   (* revision history
   hm  21. mar. 2008   rev 1.0
       original version

   hm  10. mar. 2009 rev 1.1
       real constants updated to new systax using dot

   *)
END_FUNCTION

FUNCTION "R2_ADD" : "REAL2"   // FC144, SCL
TITLE = R2_ADD
{ S7_Optimized_Access := 'FALSE' }
AUTHOR : hugo
FAMILY : R2
NAME : ADD
VERSION : 1.0
// R2_add adds a real to a double real which extends the accuracy of a real to twice as many digits
//  
// uses: REAL2 [UDT11]
   VAR_INPUT
      X : "REAL2";
      Y : Real;
   END_VAR
   VAR_TEMP
      temp : Real;
      tR2_ADD : "REAL2";
   END_VAR
BEGIN


   #temp := #X.RX;
   #tR2_ADD.RX := #Y + #X.R1 + #X.RX;
   #tR2_ADD.R1 := #temp - #tR2_ADD.RX + #Y + #X.R1;

   #R2_ADD := #tR2_ADD;

   (* revision history
   hm      20.3.2008   rev 1.0
       original version

   *)
END_FUNCTION

FUNCTION "R2_ADD2" : "REAL2"   // FC145, SCL
TITLE = R2_ADD2
{ S7_Optimized_Access := 'FALSE' }
AUTHOR : hugo
FAMILY : R2
NAME : ADD2
VERSION : 1.0
// R2_add2 adds a double precision real to a double precision real which extends the accuracy of a real to twice as many digits
//  
// uses: REAL2 [UDT11]
   VAR_INPUT
      X : "REAL2";
      Y : "REAL2";
   END_VAR
   VAR_TEMP
      tR2_ADD2 : "REAL2";
   END_VAR
BEGIN


   #tR2_ADD2.R1 := #X.R1 + #Y.R1;
   #tR2_ADD2.RX := #X.RX + #Y.RX;

   #R2_ADD2 := #tR2_ADD2;

   (* revision history
   hm      20.3.2008   rev 1.0
       original version

   *)
END_FUNCTION

FUNCTION "R2_MUL" : "REAL2"   // FC146, SCL
TITLE = R2_MUL
{ S7_Optimized_Access := 'FALSE' }
AUTHOR : hugo
FAMILY : R2
NAME : MUL
VERSION : 1.0
// R2_mul multiplies a real with a double real which extends the accuracy of a real to twice as many digits
//  
// uses: REAL2 [UDT11]
   VAR_INPUT
      X : "REAL2";
      Y : Real;
   END_VAR
   VAR_TEMP
      tR2_MUL : "REAL2";
   END_VAR
BEGIN


   #tR2_MUL.RX := #X.RX * #Y;
   #tR2_MUL.R1 := #X.R1 * #Y;

   #R2_MUL := #tR2_MUL;

   (* revision history
   hm      20.3.2008   rev 1.0
       original version

   *)
END_FUNCTION

FUNCTION "R2_SET" : "REAL2"   // FC147, SCL
TITLE = R2_SET
{ S7_Optimized_Access := 'FALSE' }
AUTHOR : hugo
FAMILY : R2
NAME : SET
VERSION : 1.1
// R2_set sets a double precision real to a single real value.
// 
// uses: REAL2 [UDT11]
   VAR_INPUT
      X : Real;
   END_VAR
   VAR_TEMP
      tR2_SET : "REAL2";
   END_VAR
BEGIN


   #tR2_SET.RX := #X;
   #tR2_SET.R1 := 0.0;

   #R2_SET := #tR2_SET;


   (* revision history
   hm  2. jun. 2008    rev 1.0
       original version

   hm  10. mar. 2009   rev 1.1
       real constants updated to new systax using dot

   *)
END_FUNCTION

// ===== PLC "Math Vektormathematik"  Unspecific CPU S7 300 =====

TYPE "VECTOR_3"
VERSION : 0.0
   STRUCT
      X : Real;
      Y : Real;
      Z : Real;
   END_STRUCT;
END_TYPE

FUNCTION "V3_ABS" : Real   // FC162, SCL
TITLE = V3_ABS
{ S7_Optimized_Access := 'FALSE' }
AUTHOR : hugo
FAMILY : MATH_V3
NAME : V3_ABS
VERSION : 1.0
// this function calculates the length of a vectors in a 3 dimensional space
// 
// uses: VECTOR_3 [UDT15]
   VAR_INPUT
      "A" : "VECTOR_3";
   END_VAR
BEGIN


   #V3_ABS := SQRT(#"A".X * #"A".X + #"A".Y * #"A".Y + #"A".Z * #"A".Z);


   (* revision history
   hm    11 dec 2007 rev 1.0
     original version

   *)
END_FUNCTION

FUNCTION "V3_ADD" : "VECTOR_3"   // FC163, SCL
TITLE = V3_ADD
{ S7_Optimized_Access := 'FALSE' }
AUTHOR : hugo
FAMILY : MATH_V3
NAME : V3_ADD
VERSION : 1.0
// this function adds two vectors in a 3 dimensional space
// 
// uses: VECTOR_3 [UDT15]
   VAR_INPUT
      "A" : "VECTOR_3";
      "B" : "VECTOR_3";
   END_VAR
BEGIN


     #V3_ADD.X := #"A".X + #"B".X;
     #V3_ADD.Y := #"A".Y + #"B".Y;
     #V3_ADD.Z := #"A".Z + #"B".Z;

     #V3_ADD := #V3_ADD;


   (* revision history
   hm    11 dec 2007 rev 1.0
     original version

   *)
END_FUNCTION

FUNCTION "V3_ANG" : Real   // FC164, SCL
TITLE = V3_ANG
{ S7_Optimized_Access := 'FALSE' }
AUTHOR : hugo
FAMILY : MATH_V3
NAME : V3_ANG
VERSION : 1.1
// this function calculates the angle between two vectors in a 3 dimensional space
// 
// uses: VECTOR_3 [UDT15]
//       V3_ABS [FC162]
//       V3_DPRO [FC165]
   VAR_INPUT
      "A" : "VECTOR_3";
      "B" : "VECTOR_3";
   END_VAR
   VAR_TEMP
      d : Real;
      temp_A : "VECTOR_3";
      temp_B : "VECTOR_3";
   END_VAR
BEGIN


   #temp_A := #"A";
   #temp_B := #"B";

   #d := "V3_ABS"(#temp_A) * "V3_ABS"(#temp_B);
   IF #d > 0.0 THEN
       #V3_ANG := ACOS(LIMIT(MN:=-1.0,IN:="V3_DPRO"(A:=#temp_A,B:=#temp_B) / #d,MX:=1.0));
   END_IF;


   (* revision history
   hm  11. dec. 2007   rev 1.0
       original version

   hm  10. mar. 2009   rev 1.1
       changed syntax of real constants to 0.0

   *)
END_FUNCTION

FUNCTION "V3_DPRO" : Real   // FC165, SCL
TITLE = V3_DPRO
{ S7_Optimized_Access := 'FALSE' }
AUTHOR : hugo
FAMILY : MATH_V3
NAME : V3_DPRO
VERSION : 1.0
// this function calculates the dot product of two vectors in 3 dimensional space
// 
// uses: VECTOR_3 [UDT15]
   VAR_INPUT
      "A" : "VECTOR_3";
      "B" : "VECTOR_3";
   END_VAR
BEGIN


     #V3_DPRO := #"A".X * #"B".X + #"A".Y * #"B".Y + #"A".Z * #"B".Z;


   (* revision history
   hm    11 dec 2007 rev 1.0
     original version

   *)
END_FUNCTION

FUNCTION "V3_NORM" : "VECTOR_3"   // FC166, SCL
TITLE = V3_NORM
{ S7_Optimized_Access := 'FALSE' }
AUTHOR : hugo
FAMILY : MATH_V3
NAME : V3_NORM
VERSION : 1.1
// this function generates a vectors with absolute length 1 from a vector A in a 3 dimensional space
// 
// uses: VECTOR_3 [UDT15]
//       V3_ABS [FC162]
//       V3_SMUL [FC170]
   VAR_INPUT
      "A" : "VECTOR_3";
   END_VAR
   VAR_TEMP
      la : Real;
      temp_A : "VECTOR_3";
      temp_V3_NORM : "VECTOR_3";
   END_VAR
BEGIN


   #temp_A := #"A";

   #la := "V3_ABS"(#temp_A);
   IF #la > 0.0 THEN
       #temp_V3_NORM := "V3_SMUL"(A:=#temp_A,M:=1.0 / #la);
   END_IF;

   #V3_NORM := #temp_V3_NORM;


   (* revision history
   hm  11 dec 2007 rev 1.0
       original version

   hm  10. mar. 2009   rev 1.1
       changed syntax of real constants to 0.0

   *)
END_FUNCTION

FUNCTION "V3_NUL" : Bool   // FC167, SCL
TITLE = V3_NUL
{ S7_Optimized_Access := 'FALSE' }
AUTHOR : hugo
FAMILY : MATH_V3
NAME : V3_NUL
VERSION : 1.1
// this function checks if a vectors in a null Vector
// 
// uses: VECTOR_3 [UDT15]
   VAR_INPUT
      "A" : "VECTOR_3";
   END_VAR
BEGIN


   #V3_NUL := #"A".X = 0.0 AND #"A".Y = 0.0 AND #"A".Z = 0.0;


   (* revision history
   hm  12 dec 2007 rev 1.0
       original version

   hm  10. mar. 2009   rev 1.1
       changed syntax of real constants to 0.0

   *)
END_FUNCTION

FUNCTION "V3_PAR" : Bool   // FC168, SCL
TITLE = V3_PAR
{ S7_Optimized_Access := 'FALSE' }
AUTHOR : hugo
FAMILY : MATH_V3
NAME : V3_PAR
VERSION : 1.1
// this function checks if two vectors in a 3 dimensional space are parallel.
// which means the two vectors have the same direction
// 
// uses: VECTOR_3 [UDT15]
//       V3_ABS [FC162]
//       V3_XPRO [FC173]
   VAR_INPUT
      "A" : "VECTOR_3";
      "B" : "VECTOR_3";
   END_VAR
   VAR_TEMP
      temp_A : "VECTOR_3";
      temp_B : "VECTOR_3";
   END_VAR
BEGIN


   #temp_A := #"A";
   #temp_B := #"B";

   #V3_PAR := "V3_ABS"("V3_XPRO"(A:=#temp_A,B:=#temp_B)) = 0.0;


   (* revision history
   hm  11 dec 2007   rev 1.0
       original version

   hm  10. mar. 2009   rev 1.1
       changed syntax of real constants to 0.0

   *)
END_FUNCTION

FUNCTION "V3_REV" : "VECTOR_3"   // FC169, SCL
TITLE = V3_REV
{ S7_Optimized_Access := 'FALSE' }
AUTHOR : hugo
FAMILY : MATH_V3
NAME : V3_REV
VERSION : 1.0
// this function reverses a vector in a 3 dimensional space
// 
// uses: VECTOR_3 [UDT15]
   VAR_INPUT
      "A" : "VECTOR_3";
   END_VAR
   VAR_TEMP
      temp_V3_REV : "VECTOR_3";
   END_VAR
BEGIN


     #temp_V3_REV.X := -#"A".X;
     #temp_V3_REV.Y := -#"A".Y;
     #temp_V3_REV.Z := -#"A".Z;

     #V3_REV := #temp_V3_REV;

   (* revision history
   hm    11 dec 2007 rev 1.0
     original version

   *)
END_FUNCTION

FUNCTION "V3_SMUL" : "VECTOR_3"   // FC170, SCL
TITLE = V3_SMUL
{ S7_Optimized_Access := 'FALSE' }
AUTHOR : hugo
FAMILY : MATH_V3
NAME : V3_SMUL
VERSION : 1.0
// this function multiplies a vectors in a 3 dimensional space with a skalar M
// 
// uses: VECTOR_3 [UDT15]
   VAR_INPUT
      "A" : "VECTOR_3";
      "M" : Real;
   END_VAR
   VAR_TEMP
      temp_V3_SMUL : "VECTOR_3";
   END_VAR
BEGIN


   #temp_V3_SMUL.X := #"A".X * #"M";
   #temp_V3_SMUL.Y := #"A".Y * #"M";
   #temp_V3_SMUL.Z := #"A".Z * #"M";

   #V3_SMUL := #temp_V3_SMUL;


   (* revision history
   hm    11 dec 2007 rev 1.0
     original version

   *)
END_FUNCTION

FUNCTION "V3_SUB" : "VECTOR_3"   // FC171, SCL
TITLE = V3_SUB
{ S7_Optimized_Access := 'FALSE' }
AUTHOR : hugo
FAMILY : MATH_V3
NAME : V3_SUB
VERSION : 1.0
// this function subtracts two vectors in a 3 dimensional space
// V3_SUB = A - B
// 
// uses: VECTOR_3 [UDT15]
   VAR_INPUT
      "A" : "VECTOR_3";
      "B" : "VECTOR_3";
   END_VAR
   VAR_TEMP
      temp_V3_SUB : "VECTOR_3";
   END_VAR
BEGIN


     #temp_V3_SUB.X := #"A".X - #"B".X;
     #temp_V3_SUB.Y := #"A".Y - #"B".Y;
     #temp_V3_SUB.Z := #"A".Z - #"B".Z;

     #V3_SUB := #temp_V3_SUB;

   (* revision history
   hm    11 dec 2007 rev 1.0
     original version

   *)
END_FUNCTION

FUNCTION "V3_XANG" : Real   // FC172, SCL
TITLE = V3_XANG
{ S7_Optimized_Access := 'FALSE' }
AUTHOR : hugo
FAMILY : MATH_V3
NAME : V3_XANG
VERSION : 1.1
// this function calculates the angle between the X-axis and a vectors in a 3 dimensional space
// 
// uses: VECTOR_3 [UDT15]
//       V3_ABS [FC162]
   VAR_INPUT
      "A" : "VECTOR_3";
   END_VAR
   VAR_TEMP
      la : Real;
      temp_A : "VECTOR_3";
   END_VAR
BEGIN


   #temp_A := #"A";

   #la := "V3_ABS"(#temp_A);
   IF #la > 0.0 THEN
       #V3_XANG := ACOS(#temp_A.X / #la);
   END_IF;


   (* revision history
   hm  11 dec 2007   rev 1.0
       original version

   hm  10. mar. 2009   rev 1.1
       changed syntax of real constants to 0.0

   *)
END_FUNCTION

FUNCTION "V3_XPRO" : "VECTOR_3"   // FC173, SCL
TITLE = V3_XPRO
{ S7_Optimized_Access := 'FALSE' }
AUTHOR : hugo
FAMILY : MATH_V3
NAME : V3_XPRO
VERSION : 1.0
// this function adds two vectors in a 3 dimensional space
// 
// uses: VECTOR_3 [UDT15]
   VAR_INPUT
      "A" : "VECTOR_3";
      "B" : "VECTOR_3";
   END_VAR
   VAR_TEMP
      temp_V3_XPRO : "VECTOR_3";
   END_VAR
BEGIN


   #temp_V3_XPRO.X := #"A".Y * #"B".Z - #"A".Z * #"B".Y;
   #temp_V3_XPRO.Y := #"A".Z * #"B".X - #"A".X * #"B".Z;
   #temp_V3_XPRO.Z := #"A".X * #"B".Y - #"A".Y * #"B".X;

   #V3_XPRO := #temp_V3_XPRO;

   (* revision history
   hm    11 dec 2007 rev 1.0
     original version

   *)
END_FUNCTION

FUNCTION "V3_YANG" : Real   // FC174, SCL
TITLE = V3_YANG
{ S7_Optimized_Access := 'FALSE' }
AUTHOR : hugo
FAMILY : MATH_V3
NAME : V3_YANG
VERSION : 1.1
// this function calculates the angle between the Y-axis and a vectors in a 3 dimensional space
// 
// uses: VECTOR_3 [UDT15]
//       V3_ABS [FC162]
   VAR_INPUT
      "A" : "VECTOR_3";
   END_VAR
   VAR_TEMP
      la : Real;
      temp_A : "VECTOR_3";
   END_VAR
BEGIN


   #temp_A := #"A";

   #la := "V3_ABS"(#temp_A);
   IF #la > 0.0 THEN
       #V3_YANG := ACOS(#temp_A.Y / #la);
   END_IF;


   (* revision history
   hm  11 dec 2007   rev 1.0
       original version

   hm  10. mar. 2009   rev 1.1
       changed syntax of real constants to 0.0

   *)
END_FUNCTION

FUNCTION "V3_ZANG" : Real   // FC175, SCL
TITLE = V3_ZANG
{ S7_Optimized_Access := 'FALSE' }
AUTHOR : hugo
FAMILY : MATH_V3
NAME : V3_ZANG
VERSION : 1.1
// this function calculates the angle between the Z-axis and a vectors in a 3 dimensional space
// 
// uses: VECTOR_3 [UDT15]
//       V3_ABS [FC162]
   VAR_INPUT
      "A" : "VECTOR_3";
   END_VAR
   VAR_TEMP
      la : Real;
      temp_A : "VECTOR_3";
   END_VAR
BEGIN


   #temp_A := #"A";

   #la := "V3_ABS"(#temp_A);
   IF #la > 0.0 THEN
       #V3_ZANG := ACOS(#temp_A.Z / #la);
   END_IF;


   (* revision history
   hm  11 dec 2007   rev 1.0
       original version

   hm  10. mar. 2009   rev 1.1
       changed syntax of real constants to 0.0

   *)
END_FUNCTION

// ===== PLC "Mathematical"  Unspecific CPU S7 300 =====

VAR_GLOBAL CONSTANT   // PLC tag table "STEP7 classic symbols"
   "PI1" : Real := 3.14159265358979323846264338327950288;
   "PI05" : Real := 1.5707963267949;
   "PI2" : Real := 6.283185307179586476;   // PI * 2
   "E_INV" : Real := 0.367879441171442;   // 1 / e
   "PI_INV" : Real := 0.318309886183791;   // 1 / PI
   "debug" : Bool := FALSE;
   "N" : Int := 0;
   "offset" : Int := 0;
   "E" : Real := 2.71828182845904523536028747135266249;   // Eulersche Konstante
   "PI" : Real := 3.14159265358979323846264338327950288;
   "offset_1" : DWord := 0;
END_VAR

TYPE "FRACTION"
VERSION : 0.0
   STRUCT
      NUMERATOR : Int;
      DENOMINATOR : Int;
   END_STRUCT;
END_TYPE

DATA_BLOCK "MATH"   // DB2
TITLE = MATH
{ S7_Optimized_Access := 'FALSE' }
AUTHOR : oscat
FAMILY : CONSTANT
NAME : DBMATH
VERSION : 1.1
   VAR
      PI : Real := 3.141593e+0;   // Kreiszahl PI
      PI2 : Real := 6.283185e+0;   // PI * 2
      PI4 : Real := 1.256637e+1;   // PI * 4
      PI05 : Real := 1.570796e+0;   // PI / 2
      PI025 : Real := 7.853982e-1;   // PI / 4
      PI_INV : Real := 3.183099e-1;   // 1 / PI
      "E" : Real := 2.718282e+0;   // Eulersche Konstante
      E_INV : Real := 3.678795e-1;   // 1 / e
      SQ2 : Real := 1.414214e+0;   // Wurzel von 2
      FACTS : Array[0..12] of DInt;
   END_VAR
BEGIN
   FACTS[0] := DINT#1;
   FACTS[1] := DINT#1;
   FACTS[2] := DINT#2;
   FACTS[3] := DINT#6;
   FACTS[4] := DINT#24;
   FACTS[5] := DINT#120;
   FACTS[6] := DINT#720;
   FACTS[7] := DINT#5040;
   FACTS[8] := DINT#40320;
   FACTS[9] := DINT#362880;
   FACTS[10] := DINT#3628800;
   FACTS[11] := DINT#39916800;
   FACTS[12] := DINT#479001600;
END_DATA_BLOCK

DATA_BLOCK "IDB_STIME"   // DB64
{ S7_Optimized_Access := 'FALSE' }
AUTHOR : dalbi
FAMILY : MEASURE
VERSION : 0.0
// stored: InstanceOfName STIME
"STIME"
BEGIN
END_DATA_BLOCK

FUNCTION_BLOCK "STIME"   // FB64, SCL
TITLE = STIME
{ S7_Optimized_Access := 'FALSE' }
AUTHOR : dalbi
FAMILY : MEASURE
NAME : STIME
VERSION : 1.4
// this function block makes sure that the timer of a siemens sps counts from 0 - 2^32-1.
   VAR_OUTPUT
      tx : DWord;
      at_tx AT tx : Array[0..31] of Bool;
   END_VAR
   VAR
      last_time : DWord;
      bit31 : Bool;
      init : Bool := TRUE;
   END_VAR
   VAR_TEMP
      TOP_SI : Struct
         EV_CLASS : Byte;
         EV_NUM : Byte;
         PRIORITY : Byte;
         NUM : Byte;
         TYP2_3 : Byte;
         TYP1 : Byte;
         ZI1 : Word;
         ZI2_3 : DWord;
      END_STRUCT;
      START_UP_SI : Struct
         EV_CLASS : Byte;
         EV_NUM : Byte;
         PRIORITY : Byte;
         NUM : Byte;
         TYP2_3 : Byte;
         TYP1 : Byte;
         ZI1 : Word;
         ZI2_3 : DWord;
      END_STRUCT;
      ERR : Int;
   END_VAR
BEGIN


   (* this FB is only necessary for siemens sps
   the siemens sps timer counts from 0 to 2^31-1 and starts at 0 sfter overrun.
   this means that the bit 31 (the highest bit ) will never be used and therefore
   a problem arises when t2 - t1 is checked.
   t2 - t1 is always valid also in an timer overrun situation where the time t1 is very high and t2 is very low.
   the result of the subtraction t2 - t1 however is still valid.
   this calculation does not work for soiemens because the highest bit is not used.

   this module stores the highest bit, changes the highest bit at every overrun occurence and stuffs ther highest bit in the output.
   the output is then used by t_plc_us and t_plc_ms.

   the correction needs and fb and not a function because the value of the highest bit has to be stored.

   do never use this function block in a codesys environment. the timer in codesys is correct and runs from 0 to 2^32-1
   *)

   (* read actual startup info *)
   (* OB1_SCAN_1  BYTE  -  B#16#01: Abschluss des Neustarts (Warmstarts)
                        -  B#16#02: Abschluss des Wiederanlaufs
                        -  B#16#03: Abschluss des freien Zyklus
                        -  B#16#04: Abschluss des Kaltstarts
                        -  B#16#05: Erster OB 1-Zyklus der neuen Master-CPU nach 
                                    Master-Reserve-Umschaltung und STOP des 
                                    bisherigen Masters *)

   #ERR := RD_SINFO (TOP_SI => #TOP_SI, START_UP_SI => #START_UP_SI);

   (* reset last_time on system startup *)
   IF #TOP_SI.EV_NUM = 1 OR #TOP_SI.EV_NUM = 2 OR #TOP_SI.EV_NUM = 4 OR NOT #init THEN 
       #last_time := 0;
       #bit31 := false;
       #init := true;
   END_IF;

   (* read the system timer *)
   #tx := DINT_TO_DWORD(T_CONV(TIME_TCK()));

   (* check for overrun *)
   IF DWORD_TO_DINT(#tx) < DWORD_TO_DINT(#last_time) THEN
       (* an overrun has occured, change the value of the highest bit *)
       #bit31 := NOT #bit31;
   END_IF;

   (* stuff the highest bit into the timer value *)
   #at_tx[7] := #bit31;

   (* remember the last system time for the next overrun check *)
   #last_time := #tx;


   (* revision history
   DA  14.9.2007 rev 1.0
     original version

   DA  24.2.2008 rev 1.1
     added self reset on system startup

   DA   2.5.2008 rev 1.2
     corect a problem running under OB35

   DA  12.3.2009 rev 1.3
     corect a problem run on different CPUs

   DA  22.12.2009 rev 1.4
     corect a problem on startup
   *)
END_FUNCTION_BLOCK

FUNCTION "DEC1" : Int   // FC52, SCL
TITLE = DEC1
{ S7_Optimized_Access := 'FALSE' }
AUTHOR : hugo
FAMILY : MATH
NAME : DEC1
VERSION : 1.1
// This is a decrement function which decrements the variable X by 1 and if 0 is reached, it begins with M again.
// _dec1(3,X) will generate 3,2,1,0,3,2,...
   VAR_INPUT
      X : Int;
      N : Int;
   END_VAR
BEGIN


   IF #X = 0 THEN
       #DEC1 := #N - 1;
   ELSE
       #DEC1 := #X - 1;
   END_IF;

   (* this is a very elegant version but 50% slower
   X := (X - 1 + N) MOD N;
   *)


   (* revision history
   hm  13. oct. 2008   rev 1.0
       original version

   hm  27. oct. 2008   rev 1.1
       added statement to return value for compatibility reasons
   *)
END_FUNCTION

FUNCTION "INC1" : Int   // FC53, SCL
TITLE = INC1
{ S7_Optimized_Access := 'FALSE' }
AUTHOR : hugo
FAMILY : MATH
NAME : INC1
VERSION : 1.2
// This is a increment function which increments the variable X by 1 and if M is reached, it begins with 0 again.
// _inc1(3,X) will generate 0,1,2,3,0,1,.....
   VAR_INPUT
      X : Int;
      N : Int;
   END_VAR
BEGIN


   IF #X >= #N - 1 THEN
       #INC1 := 0;
   ELSE
       #INC1 := #X + 1;
   END_IF;


   (* this elegant version is 50% slower
   INC1 := X := (x + 1) MOD N;
   *)



   (* revision history
   hm  13. oct. 2008   rev 1.0
       original version

   hm  22. oct. 2008   rev 1.1
       added statement to return value for compatibility reasons

   hm  23. feb. 2009   rev 1.2
       when inc1 is called with X >= N inc will continue with 0
   *)
END_FUNCTION

FUNCTION "ACOSH" : Real   // FC54, SCL
TITLE = ACOSH
{ S7_Optimized_Access := 'FALSE' }
AUTHOR : hugo
FAMILY : MATH
NAME : ACOSH
VERSION : 1.3
// this function calculates the arcus cos hyperbolicus
   VAR_INPUT
      X : Real;
   END_VAR
BEGIN



   #ACOSH := LN(SQRT(#X * #X - 1.0) + #X);


   (* revision history
   hm      12 jan 2007 rev 1.0
       original version

   hm      2. dec 2007 rev 1.1
       changed code for better performance

   hm  16. mar. 2007       rev 1.2
       changed sequence of calculations to improve performance

   hm  10. mar. 2009       rev 1.3
       real constants updated to new systax using dot

   *)
END_FUNCTION

FUNCTION "ACOTH" : Real   // FC55, SCL
TITLE = ACOTH
{ S7_Optimized_Access := 'FALSE' }
AUTHOR : hugo
FAMILY : MATH
NAME : ACOTH
VERSION : 1.2
// this function calculates the arcus cotangens hyperbolicus
   VAR_INPUT
      X : Real;
   END_VAR
BEGIN


   #ACOTH := LN((#X+1.0)/(#X-1.0))*0.5;


   (* revision history
   hm      12 jan 2007 rev 1.0
       original version

   hm      5. jan 2008 rev 1.1
       improved code for better performance

   hm  10. mar. 2009       rev 1.2
       real constants updated to new systax using dot

   *)
END_FUNCTION

FUNCTION "AGDF" : Real   // FC56, SCL
TITLE = AGDF
{ S7_Optimized_Access := 'FALSE' }
AUTHOR : hugo
FAMILY : MATH
NAME : AGDF
VERSION : 1.1
// this function calculates the inverse Gudermannian function.
   VAR_INPUT
      X : Real;
   END_VAR
BEGIN


   #AGDF := LN((1.0 + SIN(#X))/COS(#X));

   (* comment
   the current implementation gives sufficient accuracy only up to X = 1.57 or an output > 10.
   is X closer to PI/2 then the function is more and more unreliable
   *)


   (* revision history
   hm  27. apr. 2008   rev 1.0
       original version

   hm  10. mar. 2009   rev 1.1
       real constants updated to new systax using dot

   *)
END_FUNCTION

FUNCTION "ASINH" : Real   // FC57, SCL
TITLE = ASINH
{ S7_Optimized_Access := 'FALSE' }
AUTHOR : hugo
FAMILY : MATH
NAME : ASINH
VERSION : 1.3
// this function calculates the arcus sin hyperbolicus
   VAR_INPUT
      X : Real;
   END_VAR
BEGIN


   #ASINH := LN(SQRT(#X * #X + 1.0)+#X);


   (* revision history
   hm      12 jan 2007 rev 1.0
       original version

   hm      2. dec 2007 rev 1.1
       changed code for better performance

   hm      16.3. 2007      rev 1.2
       changed sequence of calculations to improve performance

   hm  10. mar. 2009       rev 1.3
       real constants updated to new systax using dot

   *)
END_FUNCTION

FUNCTION "ATAN2" : Real   // FC58, SCL
TITLE = ATAN2
{ S7_Optimized_Access := 'FALSE' }
AUTHOR : hugo
FAMILY : MATH
NAME : ATAN2
VERSION : 1.2
// this function calculates the angle in a coordinate system in rad.
   VAR_INPUT
      Y : Real;
      X : Real;
   END_VAR
BEGIN


   IF #X > 0.0 THEN
       #ATAN2 := ATAN(#Y/#X);
   ELSIF #X < 0.0 THEN
       IF #Y >= 0.0 THEN
           #ATAN2 := ATAN(#Y/#X) + "PI1";
       ELSE
           #ATAN2 := ATAN(#Y/#X) - "PI1";
       END_IF;
   ELSIF #Y > 0.0 THEN
       #ATAN2 := "PI05";
   ELSIF #Y < 0.0 THEN
       #ATAN2 := -"PI05";
   ELSE
       #ATAN2 := 0.0;
   END_IF;


   (* revision history
   hm  20.  apr. 2008  rev 1.0
       original version

   hm  18. oct. 2008   rev 1.1
       changed to use math constants

   hm  10. mar. 2009   rev 1.2
       real constants updated to new systax using dot

   *)
END_FUNCTION

FUNCTION "ATANH" : Real   // FC59, SCL
TITLE = ATANH
{ S7_Optimized_Access := 'FALSE' }
AUTHOR : hugo
FAMILY : MATH
NAME : ATANH
VERSION : 1.2
// this function calculates the arcus tangens hyperbolicus
   VAR_INPUT
      X : Real;
   END_VAR
BEGIN


   #ATANH := LN((1.0 + #X)/(1.0 - #X)) * 0.5;

   (* revision history
   hm      12 jan 2007 rev 1.0
       original version

   hm      5. jan 2008 rev 1.1
       improved code for better performance

   hm  10. mar. 2009     rev 1.2
       real constants updated to new systax using dot

   *)
END_FUNCTION

FUNCTION "BETA" : Real   // FC60, SCL
TITLE = BETA
{ S7_Optimized_Access := 'FALSE' }
AUTHOR : hugo
FAMILY : MATH
NAME : BETA
VERSION : 1.0
// this function calculates the beta function for real number > 0.
// 
// uses: GAMMA [FC84]
   VAR_INPUT
      X : Real;
      Y : Real;
   END_VAR
BEGIN


   #BETA := "GAMMA"(#X) * "GAMMA"(#Y) / "GAMMA"(#X + #Y);


   (* revision history
   hm  26. oct. 2008   rev 1.0
       original version

   *)
END_FUNCTION

FUNCTION "BINOM" : DInt   // FC61, SCL
TITLE = BINOM
{ S7_Optimized_Access := 'FALSE' }
AUTHOR : hugo
FAMILY : MATH
NAME : BINOM
VERSION : 1.0
// this FUNCTION calculates the binomialkoefficient (N over k)
   VAR_INPUT
      N : Int;
      K : Int;
   END_VAR
   VAR_TEMP
      i : Int;
      tK : Int;
      tn : Int;
   END_VAR
BEGIN


   #tK := #K;
   #tn := #N;

   IF 2 * #tK > #tn THEN
       #tK := #tn - #tK;
   END_IF;
   IF #tK > #tn THEN
       RETURN;
   ELSIF #tK = 0 OR #tK = #tn THEN
       #BINOM := 1;
   ELSIF #tK = 1 THEN
       #BINOM := #tn;
   ELSE
       #BINOM := #tn;
       #tn := #tn + 1;
       FOR #i := 2 TO #tK DO
           #BINOM := #BINOM * (#tn - #i) / #i;
       END_FOR;
   END_IF;



   (*
   binomialkoeffizient(n, k)
   1  wenn k = 0 return 1
   2  wenn 2k > n
   3      dann führe aus ergebnis \leftarrow binomialkoeffizient(n, n-k)
   4  sonst führe aus ergebnis \leftarrow n
   5          von i \leftarrow 2 bis k
   6              führe aus ergebnis \leftarrow ergebnis \cdot (n + 1 - i)
   7                        ergebnis \leftarrow ergebnis : i
   8  return ergebnis
   *)



   (* revision history
   hm  25. oct. 2008 rev 1.0
       original version


   *)
END_FUNCTION

FUNCTION "CAUCHY" : Real   // FC62, SCL
TITLE = CAUCHY
{ S7_Optimized_Access := 'FALSE' }
AUTHOR : hugo
FAMILY : MATH
NAME : CAUCHY
VERSION : 1.0
// this function calculates the Cauchy distribution function
   VAR_INPUT
      X : Real;
      T : Real;
      U : Real;
   END_VAR
   VAR_TEMP
      tmp : Real;
   END_VAR
BEGIN


   #tmp := #X - #T;
   #CAUCHY := "PI_INV" * #U / (#U*#U + #tmp*#tmp);



   (* revision hisdtory
   hm  26. oct. 2008   rev 1.0
       original version

   *)
END_FUNCTION

FUNCTION "CAUCHYCD" : Real   // FC63, SCL
TITLE = CAUCHYCD
{ S7_Optimized_Access := 'FALSE' }
AUTHOR : hugo
FAMILY : MATH
NAME : CAUCHYCD
VERSION : 1.0
// this function calculates the Cauchy distribution function
   VAR_INPUT
      X : Real;
      T : Real;
      U : Real;
   END_VAR
BEGIN


   #CAUCHYCD := 0.5 + "PI_INV" * ATAN((#X - #T) / #U);



   (* revision hisdtory
   hm  26. oct. 2008   rev 1.0
       original version

   *)
END_FUNCTION

FUNCTION "T_PLC_MS" : DWord   // FC64, SCL
TITLE = T_PLC_MS
{ S7_Optimized_Access := 'FALSE' }
AUTHOR : hugo
FAMILY : MEASURE
NAME : T_PLC_MS
VERSION : 1.2
// T_PLC_MS reads the internal PLC timer and return the time, it has the advantage to be able to set a debug mode 
// and speed up the counter to test the plc timer overrun which occurs every 50 days respectively 25 days at siemens S7
// this routine also allows to correct the behavior of s7 where the internal plc counter will not count all 32 bits.
// 
// uses: STIME [FB64],IDB_STIME [DB64]
BEGIN


   "IDB_STIME"(); 
   #T_PLC_MS := "IDB_STIME".tx; 
   (* hier muss die korrektur für step7 stattfinden
   plctime muss den vollen wertebereich von time ausnutzen:
   wenn bei step7 time -24tage bis plus 24 tage ist dann muss der timer auch beim überlauf auf -24tage springen 
   und auf keinen fall auf 0 !!!!
   für siemens muss ein weiterer fb im main eingebunden werden der sicherstellt das alle 32 bits durchgezählt werden.
   es kann nur ein fb sein den er muss sich das oberste (32te) bit merken.
   oder etwa spring s7 bei überlauf auf -24 tage????? dann wäre keine korrektur nötig.
   *)
   IF "debug" THEN
       #T_PLC_MS := DINT_TO_DWORD((DWORD_TO_DINT(SHL(IN:=#T_PLC_MS,N:="N") OR SHL(IN:=DWORD#1,N:="N"))-1) + DWORD_TO_DINT("offset_1"));
   END_IF;


   (* revision history
   hm  14.9.2007   rev 1.0
       original version

   hm  12. nov 2007    rev 1.1
       added temporaray variable tx because some compilers could not handle time() as an argument

   hm  16. nov. 2008   rev 1.2
       initialized constants with 0 for compatibility reasons
   *)
END_FUNCTION

FUNCTION "CEIL" : Int   // FC66, SCL
TITLE = CEIL
{ S7_Optimized_Access := 'FALSE' }
AUTHOR : hugo
FAMILY : MATH
NAME : CEIL
VERSION : 1.1
// This is a rounding function which returns the smallest possible integer which is greater or equal to X.
// ceil(3.14) = 4
// ceil(-3.14) = 3
   VAR_INPUT
      X : Real;
   END_VAR
BEGIN


     #CEIL := REAL_TO_INT(#X); //DINT_TO_INT(TRUNC(X));
     IF #CEIL < #X THEN
         #CEIL := #CEIL + 1;
     END_IF;

   (* code before rev 1.1
   CEIL := D_TRUNC(X);
   IF CEIL < X THEN
     ceil := ceil + 1;
   END_IF;
   *)

   (* revision history
   hm    7. feb. 2007  rev 1.0
     original version

   hm    21. mar. 2008 rev 1.1
     use REAL_TO_INT instead of trunc for compatibility reasons

   *)
END_FUNCTION

FUNCTION "CEIL2" : DInt   // FC67, SCL
TITLE = CEIL2
{ S7_Optimized_Access := 'FALSE' }
AUTHOR : hugo
FAMILY : MATH
NAME : CEIL
VERSION : 1.3
// This is a rounding function which returns the smallest possible integer which is greater or equal to X.
// ceil2(3.14) = 4
// ceil2(-3.14) = -3
   VAR_INPUT
      X : Real;
   END_VAR
BEGIN


   #CEIL2 := REAL_TO_DINT(#X);
   IF DINT_TO_REAL(#CEIL2) < #X THEN
           #CEIL2 := #CEIL2 + 1;
   END_IF;


   (* revision history
   hm  21. mar. 2008   rev 1.0
       original version

   hm  4. apr. 2008    rev 1.1
       added type conversion to avoid warnings under codesys 3.0

   hm  30. jun. 2008   rev 1.2
       added type conversion to avoid warnings under codesys 3.0

   hm  10. mar. 2009   rev 1.3
       use correct statement real_to_DINT

   *)
END_FUNCTION

FUNCTION "CMP" : Bool   // FC68, SCL
TITLE = CMP
{ S7_Optimized_Access := 'FALSE' }
AUTHOR : hugo
FAMILY : MATH
NAME : CMP
VERSION : 1.1
// this function checks two inputs x and y if they are identical with the first N digits
// example : cmp(3.141516,3.141517,6 is true.
// 
// uses: EXP10 [FC77]
//       FLOOR [FC81]
   VAR_INPUT
      X : Real;
      Y : Real;
      N : Int;
   END_VAR
   VAR_TEMP
      tmp : Real;
   END_VAR
BEGIN


   #tmp := ABS(#X);
   IF #tmp > 0.0 THEN
       #tmp := "EXP10"(INT_TO_REAL("FLOOR"((LN(#tmp)/LN(10)))-#N+1));
   ELSE
       #tmp := "EXP10"(#tmp);
   END_IF;
   #CMP := ABS(#X - #Y) < #tmp;


   (* revision history
   hm  12. mar. 2008   rev 1.0
       original version

   hm  10. mar. 2009   rev 1.1
       added type conversion for compatibility reasons
   *)
END_FUNCTION

FUNCTION "COSH" : Real   // FC69, SCL
TITLE = COSH
{ S7_Optimized_Access := 'FALSE' }
AUTHOR : hugo
FAMILY : MATH
NAME : COSH
VERSION : 1.3
// this function calculates the cos hyperbolicus
   VAR_INPUT
      X : Real;
   END_VAR
   VAR_TEMP
      t : Real;
   END_VAR
BEGIN


   #t := EXP(#X);
   #COSH := (1.0 / #t + #t) * 0.5;


   (* revision histroy
   hm  12.1.2007   rev 1.0
       original version

   hm  1.12.2007   rev 1.1
       changed code to improve performance

   hm  5. jan 2008   rev 1.2
       further performance improvement

   hm  10. mar. 2009   rev 1.3
       real constants updated to new systax using dot
   *)
END_FUNCTION

FUNCTION "COTH" : Real   // FC70, SCL
TITLE = COTH
{ S7_Optimized_Access := 'FALSE' }
AUTHOR : hugo
FAMILY : MATH
NAME : COTH
VERSION : 1.4
// this function calculates the cotangens hyperbolicus
   VAR_INPUT
      X : Real;
   END_VAR
BEGIN


   IF #X > 20.0 THEN
       #COTH :=1.0;
   ELSIF #X < -20.0 THEN
       #COTH := -1.0;
   ELSE
       #COTH := 1.0 + 2.0 / (EXP(#X * 2.0) - 1.0);
   END_IF;


   (* revision histroy
   hm      12.1.2007   rev 1.0
       original version

   hm  1.12.2007       rev 1.1
       changed code to improve performance

   hm  8. jan 2008 rev 1.2
       further improvement in performance

   hm  10. mar 2008    rev 1.3
       extended range of valid inputs to +/- INV
       changed formula for better accuracy

   hm  10. mar. 2009   rev 1.4
       real constants updated to new systax using dot
   *)
END_FUNCTION

FUNCTION "D_TRUNC" : DInt   // FC71, SCL
TITLE = D_TRUNC
{ S7_Optimized_Access := 'FALSE' }
AUTHOR : hugo
FAMILY : MATH
NAME : DTRUNC
VERSION : 1.2
// d_trunc truncates a real to a dint 1.5 will be 1 and -1.5 will be -1
// d_trunc is necessary because many systems do not offer a trunc to a dint
   VAR_INPUT
      X : Real;
   END_VAR
BEGIN


   #D_TRUNC := REAL_TO_DINT(#X);
   IF #X > 0.0 THEN
       IF DINT_TO_REAL(#D_TRUNC) > #X THEN #D_TRUNC := #D_TRUNC - 1; END_IF;
   ELSE
       IF DINT_TO_REAL(#D_TRUNC) < #X THEN #D_TRUNC := #D_TRUNC + 1; END_IF;
   END_IF;


   (* for systems that support a dint truncation this routine can be replaced by trunc() *)


   (* revision history
   hm  21. mar. 2008   rev 1.0
       original version

   hm  31. oct. 2008   rev 1.1
       optimized performance

   hm  10. mar. 2009   rev 1.2
       real constants updated to new systax using dot
   *)
END_FUNCTION

FUNCTION "DEG" : Real   // FC72, SCL
TITLE = DEG
{ S7_Optimized_Access := 'FALSE' }
AUTHOR : hugo
FAMILY : MATH
NAME : DEG
VERSION : 1.2
// this function converts degrees into Radiant
// 
// uses: MODR [FC97]
//       FLOOR2 [FC82]
   VAR_INPUT
      rad : Real;
   END_VAR
BEGIN


   #DEG := "MODR"(IN:=57.29577951308232 * #rad,DIVI:=360.0);


   (* revision history
   hm  4. aug 2006 rev 1.0
       original version

   hm 16. oct 2007 rev 1.1
       added modr statement which prohibits deg to become bigger than 360

   hm  10. mar. 2009   rev 1.2
       real constants updated to new systax using dot
   *)
END_FUNCTION

FUNCTION "DIFFER" : Bool   // FC73, SCL
TITLE = DIFFER
{ S7_Optimized_Access := 'FALSE' }
AUTHOR : hugo
FAMILY : MATH
NAME : DIFFER
VERSION : 1.1
// this function checks if in1 differs more then x from in2
// the output is true if in1 < in2 - x or in1 > in2 + X
   VAR_INPUT
      in1 : Real;
      in2 : Real;
      X : Real;
   END_VAR
BEGIN


   #DIFFER := ABS(#in1 - #in2) > #X;

   (* revision history
   hm    8. oct 2006   rev 1.0
     original version

   hm    16. mar 2008  rev 1.1
     improverd code for performance

   *)
END_FUNCTION

FUNCTION "ERF" : Real   // FC74, SCL
TITLE = ERF
{ S7_Optimized_Access := 'FALSE' }
AUTHOR : hugo
FAMILY : MATH
NAME : ERF
VERSION : 1.3
// this function calculates the erf (error) function.
// 
// uses: SGN [FC106]
   VAR_INPUT
      X : Real;
   END_VAR
   VAR_TEMP
      x2 : Real;
      ax2 : Real;
   END_VAR
BEGIN


   #x2 := #X*#X;
   #ax2 := 0.147 * #x2 + 1.0;
   #ERF := SQRT(1.0 - EXP(-#x2 * ((0.27323954473516 + #ax2)/(#ax2)))) * "SGN"(#X);


   (* revision history
   hm  7. apr. 2008    rev 1.0
       original version

   hm  30. jun. 2008   rev 1.1
       added type conversions to avoid warnings under codesys 3.0

   hm  25. oct. 2008   rev 1.2
       new code using new algorithm

   hm  10. mar. 2009   rev 1.3
       real constants updated to new systax using dot
   *)
END_FUNCTION

FUNCTION "ERFC" : Real   // FC75, SCL
TITLE = ERFC
{ S7_Optimized_Access := 'FALSE' }
AUTHOR : hugo
FAMILY : MATH
NAME : ERFC
VERSION : 1.1
// this function calculates the inverse erf (error) function.
// 
// uses: ERF [FC74]
//       SGN [FC106]
   VAR_INPUT
      X : Real;
   END_VAR
BEGIN


   #ERFC := 1.0 - "ERF"(#X);


   (* revision history
   hm  7. apr. 2008    rev 1.0
       original version

   hm  10. mar. 2009   rev 1.1
       real constants updated to new systax using dot

   *)
END_FUNCTION

FUNCTION "EVEN" : Bool   // FC76, SCL
TITLE = EVEN
{ S7_Optimized_Access := 'FALSE' }
AUTHOR : hugo
FAMILY : MATH
NAME : EVEN
VERSION : 1.2
// this function chacks an input for even value
// the output is true if the input is even.
   VAR_INPUT
      in : DInt;
   END_VAR
   VAR_TEMP
      tIN : DInt;
      _IN AT tIN : Array[0..31] of Bool;
   END_VAR
BEGIN


   #tIN := #in;
   #EVEN := NOT #_IN[24]; //EVEN := NOT in.0;

   (* revision history
   hm  1. oct 2006 rev 1.0
     ORIGINAL VERSION

   hm  01.12.2007  rev 1.1
     changed code for improved performance

   hm  21. mar. 2008 rev 1.2
     changed type of input IN from INT to DINT
   *)
END_FUNCTION

FUNCTION "EXP10" : Real   // FC77, SCL
TITLE = EXP10
{ S7_Optimized_Access := 'FALSE' }
AUTHOR : hugo
FAMILY : MATH
NAME : exp10
VERSION : 1.0
// this function calculates the exponent to the basis 10
// exp10(3) = 1000
   VAR_INPUT
      X : Real;
   END_VAR
BEGIN


     #EXP10 := EXP(#X * 2.30258509299405);

   (* revision history
   hm  2. dec 2007    rev 1.0
     original version

   *)
END_FUNCTION

FUNCTION "EXPN" : Real   // FC78, SCL
TITLE = EXPN
{ S7_Optimized_Access := 'FALSE' }
AUTHOR : hugo
FAMILY : MATH
NAME : EXPN
VERSION : 1.2
// this function calculates X to the power of N (Y = X^N) whilke N is an integer
// especially on CPU's without a floating point unit this algorythm is about 30 times faster then the IEC standard EXPT() Function
   VAR_INPUT
      X : Real;
      N : Int;
   END_VAR
   VAR_TEMP
      tempN : Int;
      _tempN AT tempN : Array[0..15] of Bool;
      tempX : Real;
      sign : Bool;
   END_VAR
BEGIN


   #tempN := #N;
   #tempX := #X;

   #sign := #_tempN[7]; //N.15
   #tempN := ABS(#tempN);
   IF #_tempN[8] THEN #EXPN := #tempX; ELSE #EXPN := 1.0; END_IF;
   #tempN := WORD_TO_INT(SHR(IN:=INT_TO_WORD(#tempN),N:=1));
   WHILE #tempN > 0 DO
      #tempX := #tempX * #tempX;
      IF #_tempN[8] THEN #EXPN := #EXPN * #tempX; END_IF;
      #tempN := WORD_TO_INT(SHR(IN:=INT_TO_WORD(#tempN),N:=1));
   END_WHILE;
   IF #sign THEN #EXPN := 1.0 / #EXPN; END_IF;


   (* revision history
   hm  4. dec 2007 rev 1.0
       original version

   hm  22. oct. 2008   rev 1.1
       optimized code

   hm  10. mar. 2009   rev 1.2
       removed nested comments
       real constants updated to new systax using dot

   *)
END_FUNCTION

FUNCTION "FACT" : DInt   // FC79, SCL
TITLE = FACT
{ S7_Optimized_Access := 'FALSE' }
AUTHOR : hugo
FAMILY : MATH
NAME : FACT
VERSION : 1.5
// this function calculates the factorial of x
// if the input is negative or higher then 12 the output will be -1.
// 
// uses: MATH [DB2]
   VAR_INPUT
      X : Int;
   END_VAR
BEGIN


   IF #X >= 0 AND #X <= 12 THEN
     #FACT := "MATH".FACTS[#X];
   ELSE
     #FACT := -1;
   END_IF;


   (* working code without array
   IF X > 12 OR X < 0 THEN
     FACT := -1;
   ELSIF X < 7 THEN
     FACT := 1;
     FOR i := 2 TO X DO
       FACT := FACT * i;
     END_FOR;
   ELSE
     FACT := 5040;
     FOR i := 8 TO X DO
       FACT := FACT * i;
     END_FOR;
   END_IF;
   *)

   (* revision history
   hm 4.3.2007   rev 1.1
     changed a critical error where while loop was indefinite.

   hm  10.12.2007  rev 1.2
     start value for i has changed to 2 for better performance

   hm  10. mar 2008  rev 1.3
     changed output of fact to dint to allow bigger values

   hm  27. oct. 2008 rev 1.4
     optimized code

   hm  26. mar. 2011 rev 1.5
     using array math.facts
   *)
END_FUNCTION

FUNCTION "FIB" : Real   // FC80, SCL
TITLE = FIB
{ S7_Optimized_Access := 'FALSE' }
AUTHOR : hugo
FAMILY : MATH
NAME : FIB
VERSION : 1.3
// this function calculates the fibonacci sequence
   VAR_INPUT
      X : Int;
   END_VAR
   VAR_TEMP
      tX : Real;
      t_1 : Real;
      t_2 : Real;
   END_VAR
BEGIN


   #t_1 := 0;
   #t_2 := 0;

   #tX := INT_TO_REAL(#X);

   IF #tX < 0 OR #tX > 46 THEN
       #FIB := -1;
   ELSIF #X < 2 THEN
       #FIB := #tX;
       RETURN;
   ELSE
       (* the fibonacci number is the sum of the two suceeding fibonaci numbers *)
       (* we store the numbers alternatively in t1 and t2 depending on pt *)
       #t_2 := 1;
       WHILE #tX > 3 DO
           #tX := #tX-2;
           #t_1 := #t_1 + #t_2;
           #t_2 := #t_1 + #t_2;
       END_WHILE;
       IF #tX > 2 THEN #t_1 := #t_1 + #t_2; END_IF;
       #FIB := #t_1 + #t_2;
   END_IF;

   (* alternative code for very big numbers

   IF X < 31 THEN
       fib := 0.4472136 * (expn(1.618034,X) - expn(-0.618034,X));
   ELSE
       fib := 0.4472133 * expn(1.618034,X);
   END_IF;

   *)

   (* revision history
   hm      27. dec 2007    rev 1.0
       original version

   hm      2. jan 2008 rev 1.1
       deleted unused variable pt

   hm      10. mar 2008    rev 1.2
       changed output to dint instead of real

   hm      26. mar. 2008   rev 1.3
       function now returns -1 for input < 0 or > 46

   *)
END_FUNCTION

FUNCTION "FLOOR" : Int   // FC81, SCL
TITLE = FLOOR
{ S7_Optimized_Access := 'FALSE' }
AUTHOR : hugo
FAMILY : MATH
NAME : FLOOR
VERSION : 1.1
// This is a rounding function which returns the biggest possible integer which is less or equal to X.
// floor(3.14) = 3
// floor(-3.14) = 4
   VAR_INPUT
      X : Real;
   END_VAR
BEGIN


   #FLOOR := REAL_TO_INT(#X);
   IF #FLOOR > #X THEN
       #FLOOR := #FLOOR - 1;
   END_IF;

   (* revision history
   hm    7. feb 2007   rev 1.0
     originlal version

   hm    21. mar. 2008 rev 1.1
     replaced trunc with real_to_int for compatibility reasons

   *)
END_FUNCTION

FUNCTION "FLOOR2" : DInt   // FC82, SCL
TITLE = FLOOR2
{ S7_Optimized_Access := 'FALSE' }
AUTHOR : hugo
FAMILY : MATH
NAME : FLOOR2
VERSION : 1.1
// This is a rounding function which returns the biggest possible integer which is less or equal to X.
// floor2(3.14) = 3
// floor2(-3.14) = -4
   VAR_INPUT
      X : Real;
   END_VAR
BEGIN


   #FLOOR2 := REAL_TO_DINT(#X);
   IF DINT_TO_REAL(#FLOOR2) > #X THEN
     #FLOOR2 := #FLOOR2 - 1;
   END_IF;

   (* revision history
   hm  21. mar. 2008   rev 1.0
       originlal version

   hm  4. apr. 2008    rev 1.1
       added type conversion to avoid warnings under codesys 3.0
   *)
END_FUNCTION

FUNCTION "FRACT" : Real   // FC83, SCL
TITLE = FRACT
{ S7_Optimized_Access := 'FALSE' }
AUTHOR : hugo
FAMILY : MATH
NAME : FRACT
VERSION : 1.3
// this function returns the fraction of a real number
// fract(3.14) = 0.14
   VAR_INPUT
      x : Real;
   END_VAR
BEGIN


   IF ABS(#x) < 2.0E9 THEN
       #FRACT := #x - DINT_TO_REAL(TRUNC(#x));
   ELSE
       #FRACT := 0.0;
   END_IF;


   (* revision history
   hm  4. aug 2006 rev 1.0
       original version

   hm  11. mar 2008    rev 1.1
       added dint_to_real for compatibility reasons
       now returns 0 for number > 2e9
       changed input to x

   hm  21. mar. 2008   rev 1.2
       use D_trunc instead of TRUNC for compatibility reasons

   hm  10. mar. 2009   rev 1.3
       real constants updated to new systax using dot

   *)
END_FUNCTION

FUNCTION "GAMMA" : Real   // FC84, SCL
TITLE = GAMMA
{ S7_Optimized_Access := 'FALSE' }
AUTHOR : hugo
FAMILY : MATH
NAME : GAMMA
VERSION : 1.3
// this function calculates the stirling function which is an approximation for the gamma function
   VAR_INPUT
      X : Real;
   END_VAR
BEGIN


   IF #X > 0 THEN
       #GAMMA := SQRT("PI2"/#X) * ("E_INV" * (#X + 1.0 / (12.0 * #X - 0.1 / #X))**#X);
   END_IF;


   (* the stirling formula is not very accurate for small values of X
   IF X >=0 THEN GAMMA := SQRT(math.PI2 * X) * EXPT(X / math.E, X); END_IF;
   *)





   (* revision history
   hm  10.12.2007  rev 1.0
       original version

   hm  18. oct. 2008   rev 1.1
       using math constants

   hm  26. oct. 2008   rev 1.2
       using new formula with better accuracy

   hm  10. mar. 2009   rev 1.3
       real constants updated to new systax using dot

   *)
END_FUNCTION

FUNCTION "GAUSS" : Real   // FC85, SCL
TITLE = GAUSS
{ S7_Optimized_Access := 'FALSE' }
AUTHOR : hugo
FAMILY : MATH
NAME : GAUSS
VERSION : 1.2
// this function calculates the gaussian density function
   VAR_INPUT
      X : Real;
      U : Real;
      SI : Real;
   END_VAR
   VAR_TEMP
      temp : Real;
      si_inv : Real;
   END_VAR
BEGIN


   #temp := #X - #U;
   #si_inv := 1.0 / #SI;
   #GAUSS := EXP(#temp * #temp * #si_inv * #si_inv * -0.5) * 0.39894228 * #si_inv;


   (* revision hisdtory
   hm  6. apr. 2008    rev 1.0
       original version

   hm  27. oct. 2008   rev 1.1
       optimized performance   

   hm  10. mar. 2009   rev 1.2
       real constants updated to new systax using dot

   *)
END_FUNCTION

FUNCTION "GAUSSCD" : Real   // FC86, SCL
TITLE = GAUSSCD
{ S7_Optimized_Access := 'FALSE' }
AUTHOR : hugo
FAMILY : MATH
NAME : GAUSSCD
VERSION : 1.1
// this function calculates the gaussian cumulative distribution function
// 
// uses: ERF [FC74]
//       SGN [FC106]
   VAR_INPUT
      X : Real;
      U : Real;
      SI : Real;
   END_VAR
BEGIN


   #GAUSSCD := ("ERF"((#X - #U)/(#SI * 1.414213562)) + 1.0) * 0.5;


   (* revision hisdtory
   hm  6. apr. 2008    rev 1.0
       original version

   hm  10. mar. 2009   rev 1.1
       real constants updated to new systax using dot

   *)
END_FUNCTION

FUNCTION "GDF" : Real   // FC87, SCL
TITLE = GDF
{ S7_Optimized_Access := 'FALSE' }
AUTHOR : hugo
FAMILY : MATH
NAME : GDF
VERSION : 1.2
// this function calculates the Gudermannian function.
   VAR_INPUT
      X : Real;
   END_VAR
BEGIN


   IF #X = 0.0 THEN
       #GDF := 0.0;
   ELSIF #X > 15.0 THEN
       #GDF := "PI05";    // Käse! math.PI05;
   ELSIF #X < -15.0 THEN
       #GDF := -"PI05";   // Käse! -math.PI05;
   ELSE
       #GDF := ATAN(EXP(#X)) * 2.0 - "PI05"; // Käse! ...math.PI05;
   END_IF;


   (* revision history
   hm  27. apr. 2008   rev 1.0
       original version

   hm  18. oct. 2008   rev 1.1
       using math constants

   hm  10. mar. 2009   rev 1.2
       real constants updated to new systax using dot

   *)
END_FUNCTION

FUNCTION "GOLD" : Real   // FC88, SCL
TITLE = GOLD
{ S7_Optimized_Access := 'FALSE' }
AUTHOR : hugo
FAMILY : MATH
NAME : GOLD
VERSION : 1.1
// this function calculates the golden function.
   VAR_INPUT
      X : Real;
   END_VAR
BEGIN


   #GOLD := (#X + SQRT(#X*#X + 4.0)) * 0.5;


   (* revision history
   hm  27. apr. 2008   rev 1.0
       original version

   hm  10. mar. 2009   rev 1.1
       real constants updated to new systax using dot

   *)
END_FUNCTION

FUNCTION "HYPOT" : Real   // FC89, SCL
TITLE = HYPOT
{ S7_Optimized_Access := 'FALSE' }
AUTHOR : hugo
FAMILY : MATH
NAME : HYPOT
VERSION : 1.0
// this function calculates the pythagorean function
   VAR_INPUT
      X : Real;
      Y : Real;
   END_VAR
BEGIN


     #HYPOT := SQRT(#X*#X + #Y*#Y);


   (* revision history
   hm  21. feb 2008  rev 1.0
     original version

   *)
END_FUNCTION

FUNCTION "INC" : Int   // FC90, SCL
TITLE = INC
{ S7_Optimized_Access := 'FALSE' }
AUTHOR : hugo
FAMILY : MATH
NAME : INC
VERSION : 1.1
// This is a increment function which increments the input X by the value D and compares the result with M.
// if the output exceeds M it will continue to count from 0 again.
   VAR_INPUT
      X : Int;
      D : Int;
      "M" : Int;
   END_VAR
BEGIN


     #INC := (#X + #D + #"M" + 1) MOD (#"M" + 1);

   (* revision history
   hm  7. feb 2007   REV 1.0
     original version

   hm  15. jan 2008  rev 1.1
     allow for neagtive increment

   *)
END_FUNCTION

FUNCTION "INC2" : Int   // FC91, SCL
TITLE = INC2
{ S7_Optimized_Access := 'FALSE' }
AUTHOR : hugo
FAMILY : MATH
NAME : INC2
VERSION : 1.0
// This function increments the input X by the value D and compares the result with U.
// if the output exceeds U it will continue to count from L again.
   VAR_INPUT
      X : Int;
      D : Int;
      L : Int;
      U : Int;
   END_VAR
   VAR_TEMP
      tmp : Int;
   END_VAR
BEGIN


   #tmp := #U - #L + 1;
   #INC2 := (#X + #D - #L + #tmp) MOD #tmp + #L;



   (* revision history
   hm  29. jun. 2008       REV 1.0
       original version


   *)
END_FUNCTION

FUNCTION "INV" : Real   // FC92, SCL
TITLE = INV
{ S7_Optimized_Access := 'FALSE' }
AUTHOR : hugo
FAMILY : MATH
NAME : INV
VERSION : 1.1
// This function calculates the result of 1 / X
   VAR_INPUT
      X : Real;
   END_VAR
BEGIN


   IF #X <> 0.0 THEN #INV := 1.0 / #X; END_IF;


   (* revision history
   hm  26. oct. 2008   rev 1.0
       original version

   hm  10. mar. 2009   rev 1.1
       real constants updated to new systax using dot

   *)
END_FUNCTION

FUNCTION "LANGEVIN" : Real   // FC93, SCL
TITLE = LANGEVIN
{ S7_Optimized_Access := 'FALSE' }
AUTHOR : hugo
FAMILY : MATH
NAME : LVIN
VERSION : 1.2
// this function calculates the langevin function
// 
// uses: COTH [FC70]
   VAR_INPUT
      X : Real;
   END_VAR
BEGIN


   IF #X = 0.0 THEN
       #LANGEVIN := 0.0;
   ELSE
       #LANGEVIN := "COTH"(#X) - 1.0 / #X;
   END_IF;


   (* revision history
   hm  10.12.2007  rev 1.0
       original version

   hm  11. mar 2008    rev 1.1
       changed formula to avoid problems when x = 0

   hm  10. mar. 2009   rev 1.2
       real constants updated to new systax using dot

   *)
END_FUNCTION

FUNCTION "MAX3" : Real   // FC94, SCL
TITLE = MAX3
{ S7_Optimized_Access := 'FALSE' }
AUTHOR : hugo
FAMILY : MATH
NAME : MAX3
VERSION : 1.1
// this function returns the highest of 3 real values
   VAR_INPUT
      in1 : Real;
      in2 : Real;
      in3 : Real;
   END_VAR
BEGIN


   #MAX3 := MAX(IN1:=MAX(IN1:=#in1,IN2:=#in2),IN2:=#in3);


   (* revision history
   hm  1.1.2007  rev 1.0
     original release

   hm  18. mar. 2011 rev 1.1
     improve performance

   *)
END_FUNCTION

FUNCTION "MIN3" : Real   // FC95, SCL
TITLE = MIN3
{ S7_Optimized_Access := 'FALSE' }
AUTHOR : hugo
FAMILY : MATH
NAME : MIN3
VERSION : 1.1
// this function returns the lowest of 3 real values
   VAR_INPUT
      in1 : Real;
      in2 : Real;
      in3 : Real;
   END_VAR
BEGIN


   #MIN3 := MIN(IN1:=MIN(IN1:=#in1,IN2:=#in2),IN2:=#in3);


   (* revision history
   hm  1.1.2007  rev 1.0
     original release

   hm  18. mar. 2011 rev 1.1
     improve performance

   *)
END_FUNCTION

FUNCTION "MID3" : Real   // FC96, SCL
TITLE = MID3
{ S7_Optimized_Access := 'FALSE' }
AUTHOR : hugo
FAMILY : MATH
NAME : MID3
VERSION : 1.2
// returns the mid value of 3 real inputs.
   VAR_INPUT
      in1 : Real;
      in2 : Real;
      in3 : Real;
   END_VAR
   VAR_TEMP
      tIN1 : Real;
      tIN2 : Real;
      tIN3 : Real;
   END_VAR
BEGIN


   #tIN1 := #in1;
   #tIN2 := #in2;
   #tIN3 := #in3;

   IF #tIN1 > #tIN2 THEN 
     #MID3 := #tIN1; 
     #tIN1 := #tIN2; 
     #tIN2 := #MID3; 
   END_IF;

   IF #tIN2 > #tIN3 THEN 
     #tIN2 := #tIN3; 
   END_IF;

   #MID3 := SEL(G:=#tIN1 > #tIN2, IN0:=#tIN2, IN1:=#tIN1);

   (*
   hm  1.1.2007  rev 1.1
     rewrote the function for better performance

   hm  18. mar. 2011 rev 1.2
     improve performance
   *)
END_FUNCTION

FUNCTION "MODR" : Real   // FC97, SCL
TITLE = MODR
{ S7_Optimized_Access := 'FALSE' }
AUTHOR : hugo
FAMILY : MATH
NAME : MODR
VERSION : 1.5
// this is a modulo funtion for real numbers
// modr(5.5,2.5) = 0.5
// 
// uses: FLOOR2 [FC82]
   VAR_INPUT
      IN : Real;
      DIVI : Real;
   END_VAR
BEGIN


   IF #DIVI = 0.0 THEN
       #MODR := 0.0;
   ELSE
       #MODR := #IN - DINT_TO_REAL("FLOOR2"(#IN / #DIVI)) * #DIVI;
   END_IF;


   (* revision history

   hm  4. aug.2006     rev 1.0